   "CH-ENV-CH-ACT" : Bool AT %I76.0, 1 s
   "CH-ENV-CH-TEMP" : Bool AT %I76.1, 1 s
   "CH-ENV-CH-TERM" : Bool AT %I76.2, 1 s
   "CH-ENV-CH-RUN" : Bool AT %I76.3, 1 s
   "BombaTorreON2" : Bool AT %M69.3, 1 s
   "HabV001(1)" : Bool AT %DB90.DBX7.6, 1 s
   "HabV002(1)" : Bool AT %DB90.DBX7.7, 1 s
   "HabV003(1)" : Bool AT %DB90.DBX8.0, 1 s
   "HabV4" : Bool AT %DB90.DBX8.1, 1 s
   "MarchaV001(1)" : Bool AT %DB90.DBX11.0, 1 s
   "MarchaV002(1)" : Bool AT %DB90.DBX11.1, 1 s
   "MarchaV003(1)" : Bool AT %DB90.DBX11.2, 1 s
   "ParadaV001(1)" : Bool AT %DB90.DBX12.5, 1 s
   "ParadaV002(1)" : Bool AT %DB90.DBX12.6, 1 s
   "ParadaV003(1)" : Bool AT %DB90.DBX12.7, 1 s
   "AnimaMenuV001" : Int AT %DB46.DBW24, 1 s
   "AnimaMenuV002" : Int AT %DB46.DBW26, 1 s
   "AnimaMenuV003" : Int AT %DB46.DBW28, 1 s
   "DeshV001" : Bool AT %DB90.DBX9.3, 1 s
   "DeshV002" : Bool AT %DB90.DBX9.4, 1 s
   "DeshV003" : Bool AT %DB90.DBX9.5, 1 s

HMI tags "CompBajaMTA"
   "HabilitaciónMC060" : Bool AT %DB74.DBX3.0, 1 s
   "HabilitaciónMC061" : Bool AT %DB74.DBX3.1, 1 s
   "HabilitaciónMC062" : Bool AT %DB74.DBX3.2, 1 s
   "HabilitaciónMC063" : Bool AT %DB74.DBX3.3, 1 s
   "HabilitaciónMC064" : Bool AT %DB74.DBX3.4, 1 s
   "HabilitaciónMC065" : Bool AT %DB74.DBX3.5, 1 s
   "DeshabilitaciónMC060" : Bool AT %DB74.DBX3.6, 1 s
   "DeshabilitaciónMC061" : Bool AT %DB74.DBX3.7, 1 s
   "DeshabilitaciónMC062" : Bool AT %DB74.DBX4.0, 1 s
   "DeshabilitaciónMC063" : Bool AT %DB74.DBX4.1, 1 s
   "DeshabilitaciónMC064" : Bool AT %DB74.DBX4.2, 1 s
   "DeshabilitaciónMC065" : Bool AT %DB74.DBX4.3, 1 s
   "MarchaMC060" : Bool AT %DB74.DBX4.4, 1 s
   "MarchaMC061" : Bool AT %DB74.DBX4.5, 1 s
   "MarchaMC062" : Bool AT %DB74.DBX4.6, 1 s
   "MarchaMC063" : Bool AT %DB74.DBX4.7, 1 s
   "MarchaMC064" : Bool AT %DB74.DBX5.0, 1 s
   "MarchaMC065" : Bool AT %DB74.DBX5.1, 1 s
   "ParadaMC060" : Bool AT %DB74.DBX5.2, 1 s
   "ParadaMC061" : Bool AT %DB74.DBX5.3, 1 s
   "ParadaMC062" : Bool AT %DB74.DBX5.4, 1 s
   "ParadaMC063" : Bool AT %DB74.DBX5.5, 1 s
   "ParadaMC064" : Bool AT %DB74.DBX5.6, 1 s
   "ParadaMC065" : Bool AT %DB74.DBX5.7, 1 s
   "AnimaMC060" : Byte AT %DB74.DBB9, 1 s
   "AnimaMC061" : Byte AT %DB74.DBB10, 1 s
   "AnimaMC062" : Byte AT %DB74.DBB11, 1 s
   "AnimaMC063" : Byte AT %DB74.DBB12, 1 s
   "AnimaMC064" : Byte AT %DB74.DBB13, 1 s
   "AnimaMC065" : Byte AT %DB74.DBB14, 1 s
   "VerMC060" : Bool, internal
   "VerMC061" : Bool, internal
   "VerMC062" : Bool, internal
   "VerMC063" : Bool, internal
   "VerMC064" : Bool, internal
   "MantM060" : Bool AT %DB74.DBX16.4, 1 s
   "MantM061" : Bool AT %DB74.DBX16.5, 1 s
   "MantM062" : Bool AT %DB74.DBX16.6, 1 s
   "MantM063" : Bool AT %DB74.DBX16.7, 1 s
   "MantM064" : Bool AT %DB74.DBX17.0, 1 s
   "AutoMC060" : Bool AT %DB93.DBX0.0, 1 s
   "AutoMC061" : Bool AT %DB93.DBX0.1, 1 s
   "AutoMC062" : Bool AT %DB93.DBX0.2, 1 s
   "AutoMC063" : Bool AT %DB93.DBX0.3, 1 s
   "AutoMC064" : Bool AT %DB93.DBX0.4, 1 s
   "SponMC060" : Real AT %DB93.DBD2, 1 s
   "SponMC061" : Real AT %DB93.DBD6, 1 s
   "SponMC062" : Real AT %DB93.DBD10, 1 s
   "SponMC063" : Real AT %DB93.DBD14, 1 s
   "SponMC064" : Real AT %DB93.DBD18, 1 s
   "SpoffMC060" : Real AT %DB93.DBD22, 1 s
   "SpoffMC061" : Real AT %DB93.DBD26, 1 s
   "SpoffMC062" : Real AT %DB93.DBD30, 1 s
   "SpoffMC063" : Real AT %DB93.DBD34, 1 s
   "SpoffMC064" : Real AT %DB93.DBD38, 1 s
   "AnimMenuMC060" : Int AT %DB93.DBW44, 1 s
   "AnimMenuMC061" : Int AT %DB93.DBW46, 1 s
   "AnimMenuMC062" : Int AT %DB93.DBW48, 1 s
   "AnimMenuMC063" : Int AT %DB93.DBW50, 1 s
   "AnimMenuMC064" : Int AT %DB93.DBW52, 1 s
   "HabilitarMC060" : Bool AT %M900.0, 1 s
   "AnularSirenaCav" : Bool AT %M600.0, 1 s
   "VerMC65" : Bool, internal

HMI tags "CompresoresAltaMTA"
   "Sop1" : Bool AT %DB124.DBX0.0, 1 s
   "Sop2" : Bool AT %DB124.DBX0.1, 1 s
   "Sop3" : Bool AT %DB124.DBX0.2, 1 s
   "ReqSop1" : Int AT %DB124.DBW8, 1 s
   "ReqSop2" : Int AT %DB124.DBW10, 1 s
   "ReqSop3" : Int AT %DB124.DBW12, 1 s
   "NinSop" : Bool AT %DB124.DBX6.0, 1 s
   "VCMP1" : Int AT %DB125.DBW2, 1 s
   "VCMP2" : Int AT %DB125.DBW4, 1 s
   "VCMP3" : Int AT %DB125.DBW6, 1 s
   "VCMP4" : Int AT %DB125.DBW8, 1 s
   "VCMP5" : Int AT %DB125.DBW10, 1 s
   "IncP1" : Bool AT %DB125.DBX15.4, 100 ms
   "IncP2" : Bool AT %DB125.DBX15.5, 100 ms
   "IncP3" : Bool AT %DB125.DBX15.6, 100 ms
   "IncP4" : Bool AT %DB125.DBX15.7, 100 ms
   "IncP5" : Bool AT %DB125.DBX16.0, 100 ms
   "DecP1" : Bool AT %DB125.DBX16.2, 1 s
   "DecP2" : Bool AT %DB125.DBX16.3, 1 s
   "DecP3" : Bool AT %DB125.DBX16.4, 1 s
   "DecP4" : Bool AT %DB125.DBX16.5, 1 s
   "DecP5" : Bool AT %DB125.DBX16.6, 1 s
   "PriRealCMP1" : Int AT %DB121.DBW16, 1 s
   "PriRealCMP2" : Int AT %DB121.DBW20, 1 s
   "PriRealCMP3" : Int AT %DB121.DBW24, 1 s
   "PriRealCMP4" : Int AT %DB121.DBW28, 1 s
   "PriRealCMP5" : Int AT %DB121.DBW32, 1 s
   "Auto1" : Bool AT %DB88.DBX10.0, 1 s
   "Auto2" : Bool AT %DB88.DBX10.1, 1 s
   "Auto3" : Bool AT %DB88.DBX10.2, 1 s
   "Auto4" : Bool AT %DB88.DBX10.3, 1 s
   "Auto5" : Bool AT %DB88.DBX10.4, 1 s
   "IndV1" : Bool AT %DB121.DBX1.5, 100 ms
   "IndV2" : Bool AT %DB121.DBX1.6, 100 ms
   "IndV3" : Bool AT %DB121.DBX1.7, 100 ms
   "IndV4" : Bool AT %DB121.DBX2.0, 100 ms
   "IndV5" : Bool AT %DB121.DBX2.1, 100 ms
   "IndR1" : Bool AT %DB121.DBX2.3, 100 ms
   "IndR2" : Bool AT %DB121.DBX2.4, 100 ms
   "IndR3" : Bool AT %DB121.DBX2.5, 100 ms
   "IndR4" : Bool AT %DB121.DBX2.6, 100 ms
   "IndR5" : Bool AT %DB121.DBX2.7, 100 ms
   "Est1" : Word AT %DB120.DBW0, 1 s
   "Est2" : Word AT %DB120.DBW2, 1 s
   "Est3" : Word AT %DB120.DBW4, 1 s
   "Est4" : Word AT %DB120.DBW6, 1 s
   "Est5" : Word AT %DB120.DBW8, 1 s
   "LimSUP1" : Real AT %DB122.DBD0, 1 s
   "LimSUP2" : Real AT %DB122.DBD4, 1 s
   "LimSUP3" : Real AT %DB122.DBD8, 1 s
   "LimSUP4" : Real AT %DB122.DBD12, 1 s
   "LimSUP5" : Real AT %DB122.DBD16, 1 s
   "LimINF1" : Real AT %DB122.DBD24, 1 s
   "LimINF2" : Real AT %DB122.DBD28, 1 s
   "LimINF3" : Real AT %DB122.DBD32, 1 s
   "LimINF4" : Real AT %DB122.DBD36, 1 s
   "LimINF5" : Real AT %DB122.DBD40, 1 s
   "PresMaX" : Real AT %DB122.DBD56, 1 s
   "Delta" : Real AT %DB122.DBD48, 1 s
   "Hist" : Real AT %DB122.DBD52, 1 s
   "CompReq" : Int AT %DB121.DBW4, 1 s
   "CompReqINI" : Int AT %DB124.DBW14, 1 s
   "AnimMenuMC001" : Int AT %DB135.DBW0, 1 s
   "AnimMenuMC002" : Int AT %DB135.DBW2, 1 s
   "AnimMenuMC003" : Int AT %DB135.DBW4, 1 s
   "AnimMenuMC004" : Int AT %DB135.DBW6, 1 s
   "AnimMenuMC005" : Int AT %DB135.DBW8, 1 s
   "SPON1" : Real AT %DB135.DBD12, 1 s
   "SPON2" : Real AT %DB135.DBD16, 1 s
   "SPON3" : Real AT %DB135.DBD20, 1 s
   "SPON4" : Real AT %DB135.DBD24, 1 s
   "SPON5" : Real AT %DB135.DBD28, 1 s
   "SPOFF1" : Real AT %DB135.DBD36, 1 s
   "SPOFF2" : Real AT %DB135.DBD40, 1 s
   "SPOFF3" : Real AT %DB135.DBD44, 1 s
   "SPOFF4" : Real AT %DB135.DBD48, 1 s
   "SPOFF5" : Real AT %DB135.DBD52, 1 s
   "MantMC001" : Bool AT %DB135.DBX60.0, 1 s
   "MantMC002" : Bool AT %DB135.DBX60.1, 1 s
   "MantMC003" : Bool AT %DB135.DBX60.2, 1 s
   "MantMC004" : Bool AT %DB135.DBX60.3, 1 s
   "MantMC005" : Bool AT %DB135.DBX60.4, 1 s
   "IndVparp1" : Bool AT %DB121.DBX70.0, 1 s
   "IndVparp2" : Bool AT %DB121.DBX70.1, 1 s
   "IndVparp3" : Bool AT %DB121.DBX70.2, 1 s
   "IndVparp4" : Bool AT %DB121.DBX70.3, 1 s
   "IndVparp5" : Bool AT %DB121.DBX70.4, 1 s
   "TiempoenVacío" : Int AT %DB123.DBW4, 1 s
   "TiemposinReq" : Int AT %DB123.DBW10, 1 s
   "TiempoSop" : Int AT %DB124.DBW4, 1 s
   "HistCRT" : Real AT %DB122.DBD60, 1 s
   "LimINFCRT" : Real AT %DB122.DBD68, 1 s
   "LimSUPCRT" : Real AT %DB122.DBD64, 1 s
   "PanMCH1" : Bool AT %DB88.DBX6.0, 1 s
   "PanMCH2" : Bool AT %DB88.DBX6.1, 1 s
   "PanMCH3" : Bool AT %DB88.DBX6.2, 1 s
   "PanMCH4" : Bool AT %DB88.DBX6.3, 1 s
   "PanMCH5" : Bool AT %DB88.DBX6.4, 1 s
   "MarchaMC001" : Bool AT %DB135.DBX61.4, 1 s
   "MarchaMC002" : Bool AT %DB135.DBX61.5, 1 s
   "MarchaMC003" : Bool AT %DB135.DBX61.6, 1 s
   "MarchaMC004" : Bool AT %DB135.DBX61.7, 1 s
   "MarchaMC005" : Bool AT %DB135.DBX62.0, 1 s
   "ParadaMC001" : Bool AT %DB135.DBX62.2, 1 s
   "ParadaMC002" : Bool AT %DB135.DBX62.3, 1 s
   "ParadaMC003" : Bool AT %DB135.DBX62.4, 1 s
   "ParadaMC004" : Bool AT %DB135.DBX62.5, 1 s
   "ParadaMC005" : Bool AT %DB135.DBX62.6, 1 s
   "AnimMotorMC001" : Byte AT %DB46.DBB40, 1 s
   "AnimMotorMC002" : Byte AT %DB46.DBB41, 1 s
   "AnimMotorMC003" : Byte AT %DB46.DBB42, 1 s
   "AnimMotorMC004" : Byte AT %DB46.DBB43, 1 s
   "AnimMotorMC005" : Byte AT %DB46.DBB44, 1 s
   "EV1" : Bool AT %Q2.0, 1 s
   "EV2" : Bool AT %Q2.1, 1 s
   "EV3" : Bool AT %Q2.2, 1 s
   "EV4" : Bool AT %Q2.3, 1 s
   "EV5" : Bool AT %Q2.4, 1 s
   "HORAS1" : DInt AT %DB73.DBD0, 1 s
   "HORAS2" : DInt AT %DB73.DBD4, 1 s
   "HORAS3" : DInt AT %DB73.DBD8, 1 s
   "HORAS4" : DInt AT %DB73.DBD12, 1 s
   "HORAS5" : DInt AT %DB73.DBD16, 1 s
   "MIN1" : Int AT %DB73.DBW24, 1 s
   "MIN2" : Int AT %DB73.DBW26, 1 s
   "MIN3" : Int AT %DB73.DBW28, 1 s
   "MIN4" : Int AT %DB73.DBW30, 1 s
   "MIN5" : Int AT %DB73.DBW32, 1 s
   "MarchaOK1" : Bool AT %DB135.DBX60.6, 1 s
   "MarchaOK2" : Bool AT %DB135.DBX60.7, 1 s
   "MarchaOK3" : Bool AT %DB135.DBX61.0, 1 s
   "MarchaOK4" : Bool AT %DB135.DBX61.1, 1 s
   "MarchaOK5" : Bool AT %DB135.DBX61.2, 1 s
   "ForzarMarcha1" : Bool AT %DB136.DBX0.0, 1 s
   "ForzarMarcha2" : Bool AT %DB136.DBX0.1, 1 s
   "ForzarMarcha3" : Bool AT %DB136.DBX0.2, 1 s
   "ForzarMarcha4" : Bool AT %DB136.DBX0.3, 1 s
   "ForzarMarcha5" : Bool AT %DB136.DBX0.4, 1 s
   "ForzarParada1" : Bool AT %DB136.DBX0.6, 1 s
   "ForzarParada2" : Bool AT %DB136.DBX0.7, 1 s
   "ForzarParada3" : Bool AT %DB136.DBX1.0, 1 s
   "ForzarParada4" : Bool AT %DB136.DBX1.1, 1 s
   "ForzarParada5" : Bool AT %DB136.DBX1.2, 1 s
   "SPONF1" : Real AT %DB136.DBD4, 1 s
   "SPONF2" : Real AT %DB136.DBD8, 1 s
   "SPONF3" : Real AT %DB136.DBD12, 1 s
   "SPONF4" : Real AT %DB136.DBD16, 1 s
   "SPONF5" : Real AT %DB136.DBD20, 1 s
   "SPOFFF1" : Real AT %DB136.DBD28, 1 s
   "SPOFFF2" : Real AT %DB136.DBD32, 1 s
   "SPOFFF3" : Real AT %DB136.DBD36, 1 s
   "SPOFFF4" : Real AT %DB136.DBD40, 1 s
   "SPOFFF5" : Real AT %DB136.DBD44, 1 s
   "ForzandoMarcha1" : Bool AT %DB136.DBX1.4, 1 s
   "ForzandoMarcha2" : Bool AT %DB136.DBX1.5, 1 s
   "ForzandoMarcha3" : Bool AT %DB136.DBX1.6, 1 s
   "ForzandoMarcha4" : Bool AT %DB136.DBX1.7, 1 s
   "ForzandoMarcha5" : Bool AT %DB136.DBX2.0, 1 s
   "MediaCargaBellis" : Bool AT %DB135.DBX63.0, 1 s
   "SPONF3b" : Real AT %DB136.DBD52, 1 s
   "SPOFFF3b" : Real AT %DB136.DBD56, 1 s
   "EV3b" : Bool AT %Q3.2, 1 s
   "TiempoMaxBellismedia" : Int AT %DB63.DBW4, 1 s
   "Est6" : Int AT %DB120.DBW10, 1 s
   "PriRealCMP6" : Int AT %DB121.DBW36, 1 s
   "IndV6" : Bool AT %DB121.DBX2.2, 1 s

HMI tags "IluminaciónMTA"
   "TiempoIluminación" : Word AT %DB87.DBW0, 1 s
   "EncendidoPanel" : Bool AT %DB87.DBX2.0, 1 s
   "ApagadoPanel" : Bool AT %DB87.DBX2.1, 1 s
   "ON" : Bool AT %DB87.DBX2.2, 1 s
   "MantenerON" : Bool AT %DB87.DBX2.3, 1 s
   "AlarmaBoosters" : Bool AT %M330.4, 1 s

HMI tags "SecadoresAltaMTA"
   "AnimaMS050" : Byte AT %DB81.DBB6, 1 s
   "AnimaMS051" : Byte AT %DB81.DBB7, 1 s
   "AnimaMS052" : Byte AT %DB81.DBB8, 1 s
   "AnimaMS053" : Byte AT %DB81.DBB9, 1 s
   "DeshabilitaciónMS050" : Bool AT %DB81.DBX2.4, 1 s
   "DeshabilitaciónMS051" : Bool AT %DB81.DBX2.5, 1 s
   "DeshabilitaciónMS052" : Bool AT %DB81.DBX2.6, 1 s
   "DeshabilitaciónMS053" : Bool AT %DB81.DBX2.7, 1 s
   "HabilitaciónMS050" : Bool AT %DB81.DBX2.0, 1 s
   "HabilitaciónMS051" : Bool AT %DB81.DBX2.1, 1 s
   "HabilitaciónMS052" : Bool AT %DB81.DBX2.2, 1 s
   "HabilitaciónMS053" : Bool AT %DB81.DBX2.3, 1 s
   "MantMS050" : Bool AT %DB81.DBX11.0, 1 s
   "MantMS051" : Bool AT %DB81.DBX11.1, 1 s
   "MantMS052" : Bool AT %DB81.DBX11.2, 1 s
   "MantMS053" : Bool AT %DB81.DBX11.3, 1 s
   "MarchaMS050" : Bool AT %DB81.DBX3.0, 1 s
   "MarchaMS051" : Bool AT %DB81.DBX3.1, 1 s
   "MarchaMS052" : Bool AT %DB81.DBX3.2, 1 s
   "MarchaMS053" : Bool AT %DB81.DBX3.3, 1 s
   "ParadaMS050" : Bool AT %DB81.DBX3.4, 1 s
   "ParadaMS051" : Bool AT %DB81.DBX3.5, 1 s
   "ParadaMS052" : Bool AT %DB81.DBX3.6, 1 s
   "ParadaMS053" : Bool AT %DB81.DBX3.7, 1 s
   "AnimaMenuMS050" : Int AT %DB46.DBW14, 1 s
   "AnimaMenuMS051" : Int AT %DB46.DBW16, 1 s
   "AnimaMenuMS052" : Int AT %DB46.DBW18, 1 s
   "AnimaMenuMS053" : Int AT %DB46.DBW20, 1 s
   "Enc1MS050" : Int AT %DB81.DBW12, 1 s
   "Enc2MS050" : Int AT %DB81.DBW14, 1 s
   "Enc1MS051" : Int AT %DB81.DBW16, 1 s
   "Enc2MS051" : Int AT %DB81.DBW18, 1 s
   "Enc1MS052" : Int AT %DB81.DBW20, 1 s
   "Enc2MS052" : Int AT %DB81.DBW22, 1 s
   "Enc1MS053" : Int AT %DB81.DBW24, 1 s
   "Enc2MS053" : Int AT %DB81.DBW26, 1 s
   "AutoMS050" : Bool AT %DB81.DBX28.0, 1 s
   "AutoMS051" : Bool AT %DB81.DBX28.1, 1 s
   "AutoMS052" : Bool AT %DB81.DBX28.2, 1 s
   "AutoMS053" : Bool AT %DB81.DBX28.3, 1 s

HMI tags "SecadoresBaja"
   "AnimaMS054" : Byte AT %DB46.DBB30, 1 s
   "AnimaMS055" : Byte AT %DB46.DBB31, 1 s
   "DeshabilitaciónMS054" : Bool AT %DB49.DBX1.2, 1 s
   "DeshabilitaciónMS055" : Bool AT %DB49.DBX1.3, 1 s
   "HabilitaciónMS054" : Bool AT %DB49.DBX1.0, 1 s
   "HabilitaciónMS055" : Bool AT %DB49.DBX1.1, 1 s
   "MarchaMS054" : Bool AT %DB49.DBX1.4, 1 s
   "MarchaMS055" : Bool AT %DB49.DBX1.5, 1 s
   "ParadaMS054" : Bool AT %DB49.DBX1.6, 1 s
   "ParadaMS055" : Bool AT %DB49.DBX1.7, 1 s
   "MantMS054" : Bool AT %DB49.DBX5.4, 1 s
   "MantMS055" : Bool AT %DB49.DBX5.5, 1 s

HMI tags "SENTRON PAC 3200"
   "Tension Fase R" : Float AT %MW1, 1 s
   "Tension fase S" : Float AT %MW3, 1 s
   "Tension Fase T" : Float AT %MW5, 1 s
   "Tension Linea RS" : Float AT %MW7, 1 s
   "Tension Linea ST" : Float AT %MW9, 1 s
   "Tension Linea TR" : Float AT %MW11, 1 s
   "Corriente fase R" : Float AT %MW13, 1 s
   "Corriente Fase S" : Float AT %MW15, 1 s
   "Corriente Fase T" : Float AT %MW17, 1 s
   "Pot.Apa R" : Float AT %MW19, 1 s
   "Pot.Apa S" : Float AT %MW21, 1 s
   "Pot.Apa T" : Float AT %MW23, 1 s
   "Pot.Act R" : Float AT %MW25, 1 s
   "Pot.Act S" : Float AT %MW27, 1 s
   "Pot.Act T" : Float AT %MW29, 1 s
   "Pot.ReAct R" : Float AT %MW31, 1 s
   "Pot.ReAct S" : Float AT %MW33, 1 s
   "Pot.ReAct T" : Float AT %MW35, 1 s
   "Coseno R" : Float AT %MW37, 1 s
   "Coseno S" : Float AT %MW39, 1 s
   "Coseno T" : Float AT %MW41, 1 s
   "THD-R TensionFase R" : Float AT %MW43, 1 s
   "THD-R Tension Fase S" : Float AT %MW45, 1 s
   "THD-R Tension Fase T" : Float AT %MW47, 1 s
   "THD-R Corriente Fase R" : Float AT %MW49, 1 s
   "THD-R Corriente Fase S" : Float AT %MW51, 1 s
   "THD-R Corriente Fase T" : Float AT %MW53, 1 s
   "Frecuencia" : Float AT %MW55, 1 s
   "Tension Media Fase" : Float AT %MW57, 1 s
   "Tension Media de Linea" : Float AT %MW59, 1 s
   "Corriente Media" : Float AT %MW61, 1 s
   "Pot Apa Total" : Float AT %MW63, 1 s
   "Pot Act Total" : Float AT %MW65, 1 s
   "Pot ReAct Total" : Float AT %MW67, 1 s
   "coseno Total" : Float AT %MW69, 1 s
   "desbalance de tension" : Float AT %MW71, 1 s
   "desbalance de corriente" : Float AT %MW73, 1 s
   "Tension Maxima R" : Float AT %MW75, 1 s
   "Tension Maxima S" : Float AT %MW77, 1 s
   "Tension Maxima T" : Float AT %MW79, 1 s
   "Tension Maxima RS" : Float AT %MW81, 1 s
   "Tension Maxima ST" : Float AT %MW83, 1 s
   "Tension Maxima TR" : Float AT %MW85, 1 s
   "Corriente Maxima R" : Float AT %MW87, 1 s
   "Corriente Maxima S" : Float AT %MW89, 1 s
   "Corriente Maxima T" : Float AT %MW91, 1 s

HMI tags "TorresCav-MTA"
   "AnimaMV030" : Byte AT %DB46.DBB36, 1 s
   "AnimaMV031" : Byte AT %DB46.DBB37, 1 s
   "AnimaMP014" : Byte AT %DB46.DBB38, 1 s
   "AnimaMP015" : Byte AT %DB46.DBB39, 1 s
   "DeshabilitaciónMV030" : Bool AT %DB21.DBX2.4, 1 s
   "DeshabilitaciónMV031" : Bool AT %DB21.DBX2.5, 1 s
   "DeshabilitaciónMP014" : Bool AT %DB21.DBX2.6, 1 s
   "DeshabilitaciónMP015" : Bool AT %DB21.DBX2.7, 1 s
   "HabilitaciónMV030" : Bool AT %DB21.DBX2.0, 1 s
   "HabilitaciónMV031" : Bool AT %DB21.DBX2.1, 1 s
   "HabilitaciónMP014" : Bool AT %DB21.DBX2.2, 1 s
   "HabilitaciónMP015" : Bool AT %DB21.DBX2.3, 1 s
   "MantMV030" : Bool AT %DB21.DBX10.0, 1 s
   "MantMV031" : Bool AT %DB21.DBX10.1, 1 s
   "MantMP014" : Bool AT %DB21.DBX10.2, 1 s
   "MantMP015" : Bool AT %DB21.DBX10.3, 1 s
   "MarchaMV030" : Bool AT %DB21.DBX3.0, 1 s
   "MarchaMV031" : Bool AT %DB21.DBX3.1, 1 s
   "MarchaMP014" : Bool AT %DB21.DBX3.2, 1 s
   "MarchaMP015" : Bool AT %DB21.DBX3.3, 1 s
   "ParadaMV030" : Bool AT %DB21.DBX3.4, 1 s
   "ParadaMV031" : Bool AT %DB21.DBX3.5, 1 s
   "ParadaMP014" : Bool AT %DB21.DBX3.6, 1 s
   "ParadaMP015" : Bool AT %DB21.DBX3.7, 1 s
   "MenuV030" : Int AT %DB46.DBW32, 1 s
   "MenuV031" : Int AT %DB46.DBW34, 1 s

discrete alarms
   1: 'Falla Conexión con sensor de Temperatura torres de Cavaleto', class MTA, trigger "Rec13" bit 9
   2: 'Falla Conexión con sensor de Temperatura torres de Chillers', class MTA, trigger "Rec13" bit 10
   3: 'Falla Conexión con sensor de Presión de ALTA', class MTA, trigger "Rec13" bit 11
   4: 'Falla Conexión con sensor de Presión de ALTA redundante', class MTA, trigger "Rec13" bit 12
   5: 'Falla Conexión con sensor de Presión de Baja', class MTA, trigger "Rec13" bit 13
   6: 'Falla Presión de Alta en Límite Mínimo', class MTA, trigger "Rec13" bit 14
   7: 'Falla Presión de Alta en demasiado Baja', class MTA, trigger "Rec13" bit 15
   8: 'Falla Presión de Alta en demasiado Alta', class MTA, trigger "Rec14" bit 8
   9: 'Falla Presión de Alta en Límite Máximo', class MTA, trigger "Rec14" bit 9
   10: 'Falla Presión de Baja en Límite Mínimo', class MTA, trigger "Rec14" bit 10
   11: 'Falla Presión de Baja en demasiado Baja', class MTA, trigger "Rec14" bit 11
   12: 'Falla Presión de Baja en demasiado Alta', class MTA, trigger "Rec14" bit 12
   13: 'Falla Contactor - MS050 - Secador de Alta ABC1', class MTA, trigger "Rec6" bit 8
   14: 'Falla Guardamotor - MS051 - Secador de Alta ABC3', class MTA, trigger "Rec6" bit 9
   15: 'Falla Presión de Baja en Límite Máximo', class MTA, trigger "Rec14" bit 13
   16: 'Falla en chiller de envasado chico', class MTA, trigger "Rec14" bit 14
   17: 'Falla en chiller de soplado chico', class MTA, trigger "Rec14" bit 15
   18: 'El Compresor ABC2 alcanzó la máxima cantidad de horas sin mantenimiento #1', class MTA, trigger "Rec15" bit 8
   19: 'El Compresor ABC3 alcanzó la máxima cantidad de horas sin mantenimiento #1', class MTA, trigger "Rec15" bit 9
   20: 'El Compresor Bellis alcanzó la máxima cantidad de horas sin mantenimiento #1', class MTA, trigger "Rec15" bit 10
   21: 'El Compresor ABC4 alcanzó la máxima cantidad de horas sin mantenimiento #1', class MTA, trigger "Rec15" bit 11
   22: 'El Compresor ABC5 alcanzó la máxima cantidad de horas sin mantenimiento #1', class MTA, trigger "Rec15" bit 12
   23: 'Falla algún contactor en Booster 1', class MTA, trigger "Rec15" bit 13
   24: 'Falla algún guardamotor en Booster 1', class MTA, trigger "Rec15" bit 14
   25: 'Presión Alta en Booster', class MTA, trigger "Rec15" bit 15
   26: 'Falla algún contactor en Booster 2', class MTA, trigger "Rec16" bit 8
   27: 'Falla algún guardamotor en Booster 2', class MTA, trigger "Rec16" bit 9
   28: 'Error lectura analógica Presión Boosters', class MTA, trigger "Rec16" bit 10
   29: 'Bombas Torres de Agua Cavaleto detenidas por falla en Flujostato', class MTA, trigger "Rec16" bit 11
   30: 'Ventiladores Torres de Agua Cavaleto detenidas por falla en Flujostato', class MTA, trigger "Rec16" bit 12
   31: 'Ninguna Bomba Torres de Agua Cabaleto en Marcha', class MTA, trigger "Rec16" bit 13
   32: 'Compresores Alta Detenidos por Flujostato Torres de Agua Cabaleto', class MTA, trigger "Rec16" bit 14
   33: 'Compresores Alta Detenidos por Ninguna Bomba en Marcha en Torres de Agua Cabaleto', class MTA, trigger "Rec16" bit 15
   50: 'Falla Contactor - MS051 - Secador de Alta ABC3', class MTA, trigger "Rec6" bit 10
   53: 'Falla Guardamotor - MS052 - Secador de Alta ABC2', class MTA, trigger "Rec6" bit 11
   66: 'Falla Guardamotor MS054 - Secador de Baja SULLAIR 1', class MTA, trigger "Rec7" bit 8
   67: 'Falla Contactor MS054 - Secador de Baja SULLAIR 1', class MTA, trigger "Rec7" bit 9
   68: 'Falla Guardamotor MS055 - Secador de Baja SULLAIR 2', class MTA, trigger "Rec7" bit 10
   69: 'Falla Contactor MS055 - Secador de Baja SULLAIR 2', class MTA, trigger "Rec7" bit 11
   70: 'Falla Guardamotor - MV030 - Ventilador 2 Torres de enfriamiento Cavaleto', class MTA, trigger "Rec7" bit 12
   71: 'Falla Contactor - MV030 - Ventilador 2 Torres de enfriamiento Cavaleto', class MTA, trigger "Rec7" bit 13
   72: 'Falla Guardamotor - MV031 - Ventilador 1 Torres de enfriamiento Cavaleto', class MTA, trigger "Rec7" bit 14
   73: 'Falla Contactor - MV031 - Ventilador 1 Torres de enfriamiento Cavaleto', class MTA, trigger "Rec7" bit 15
   74: 'Falla Guardamotor - MP014 - Bomba 1 Torres de enfriamiento Cavaleto', class MTA, trigger "Rec8" bit 8
   75: 'Falla Contactor - MP014 - Bomba 1 Torres de enfriamiento Cavaleto', class MTA, trigger "Rec8" bit 9
   76: 'Falla Guardamotor - MP015 - Bomba 2 Torres de enfriamiento Cavaleto', class MTA, trigger "Rec8" bit 10
   77: 'Falla Contactor - MP015 - Bomba 2 Torres de enfriamiento Cavaleto', class MTA, trigger "Rec8" bit 11
   78: 'Falla Guardamotor - MC001 - Compresor de Alta ABC2', class MTA, trigger "Rec8" bit 12
   79: 'Falla Contactor - MC001 - Compresor de Alta ABC2', class MTA, trigger "Rec8" bit 13
   80: 'Falla Guardamotor - MC002 - Compresor de Alta ABC3', class MTA, trigger "Rec8" bit 14
   81: 'Falla Contactor - MC002 - Compresor de Alta ABC3', class MTA, trigger "Rec8" bit 15
   82: 'Falla Guardamotor - MC003 - Compresor de Alta BELLIS', class MTA, trigger "Rec9" bit 8
   83: 'Falla Contactor - MC003 - Compresor de Alta BELLIS', class MTA, trigger "Rec9" bit 9
   87: 'Falla Contactor - MS052 - Secador de Alta ABC2', class MTA, trigger "Rec6" bit 12
   88: 'Falla Guardamotor - MS053 - Secador de Alta FARGON', class MTA, trigger "Rec6" bit 13
   89: 'Falla Contactor - MS053 - Secador de Alta FARGON', class MTA, trigger "Rec6" bit 14
   90: 'Falla Presostato Chillers', class MTA, trigger "Rec6" bit 15
   91: 'Falla Guardamotor - MC004 - Compresor de Alta ABC4', class MTA, trigger "Rec9" bit 10
   92: 'Falla Contactor - MC004 - Compresor de Alta ABC4', class MTA, trigger "Rec9" bit 11
   93: 'Falla Guardamotor - MC005 - Compresor de Alta ABC5', class MTA, trigger "Rec9" bit 12
   94: 'Falla Contactor - MC005 - Compresor de Alta ABC5', class MTA, trigger "Rec9" bit 13
   95: 'Falla Flujostato Torres Caveleto', class MTA, trigger "Rec9" bit 14
   96: 'Falla Compresor ABC2 Baja Presion de Aceite', class MTA, trigger "Rec9" bit 15
   97: 'Falla Compresor ABC2 Baja Presion de Agua', class MTA, trigger "Rec10" bit 8
   98: 'Falla Compresor ABC2 Alta Temperatura de Aire', class MTA, trigger "Rec10" bit 9
   99: 'Falla Compresor ABC2 Alta Temperatura de agua', class MTA, trigger "Rec10" bit 10
   100: 'Falla Compresor ABC3 Baja Presion de Aceite', class MTA, trigger "Rec10" bit 11
   101: 'Falla Compresor ABC3 Baja Presion de Agua', class MTA, trigger "Rec10" bit 12
   102: 'Falla Compresor ABC3 Alta Temperatura de Aire', class MTA, trigger "Rec10" bit 13
   103: 'Falla Compresor ABC3 Alta Temperatura de agua', class MTA, trigger "Rec10" bit 14
   104: 'Falla Compresor ABC4 Baja Presion de Aceite', class MTA, trigger "Rec10" bit 15
   105: 'Falla Compresor ABC4 Alta Temperatura de Aire', class MTA, trigger "Rec11" bit 8
   106: 'Falla Compresor ABC4 Alta Temperatura de Aire', class MTA, trigger "Rec11" bit 9
   107: 'Falla Compresor ABC4 Alta Temperatura de agua', class MTA, trigger "Rec11" bit 10
   108: 'Falla Compresor ABC5 Baja Presion de Aceite', class MTA, trigger "Rec11" bit 11
   109: 'Falla Compresor ABC5 Alta Temperatura de Aire', class MTA, trigger "Rec11" bit 12
   110: 'Falla Compresor ABC5 Alta Temperatura de Aire', class MTA, trigger "Rec11" bit 13
   111: 'Falla Compresor ABC5 Alta Temperatura de agua', class MTA, trigger "Rec11" bit 14
   112: 'Falla Compresor Bellis & MHW28 Baja Presion Aceite', class MTA, trigger "Rec11" bit 15
   113: 'Falla Compresor Bellis & MHW28 Baja Presion de Agua', class MTA, trigger "Rec12" bit 8
   114: 'Falla Compresor Bellis & MHW28 Alta temperatura de Aire', class MTA, trigger "Rec12" bit 9
   115: 'Falla Compresor Bellis & MHW28 Alta temperatura de Agua', class MTA, trigger "Rec12" bit 10
   116: 'Falla Compresor Bellis & MHW28 Falla de Flujostato', class MTA, trigger "Rec12" bit 11
   117: 'Compresor ABC2 Requiere Marcha', class MTA, trigger "Rec12" bit 12
   118: 'Compresor ABC3 Requiere Marcha', class MTA, trigger "Rec12" bit 13
   119: 'Compresor Bellis Requiere Marcha', class MTA, trigger "Rec12" bit 14
   120: 'Compresor ABC4 Requiere Marcha', class MTA, trigger "Rec12" bit 15
   121: 'Compresor ABC5 Requiere Marcha', class MTA, trigger "Rec13" bit 8
   125: 'Falla Contactor - V001 - Ventilador 1 Torres de enfriamiento Chillers', class MTA, trigger "Rec4" bit 8
   126: 'Falla Guardamotor - V001 - Ventilador 1 Torres de enfriamiento Chillers', class MTA, trigger "Rec3" bit 15
   127: 'Falla Guardamotor - V003 - Ventilador 3 Torres de enfriamiento Chillers', class MTA, trigger "Rec4" bit 11
   128: 'Falla Contactor - V002 - Ventilador 2 Torres de enfriamiento Chillers', class MTA, trigger "Rec4" bit 10
   129: 'Falla Guardamotor - V002 - Ventilador 2 Torres de enfriamiento Chillers', class MTA, trigger "Rec4" bit 9
   130: 'Falla Guardamotor - MP018 - Bomba 1 Torres de enfriamiento Chillers', class MTA, trigger "Rec3" bit 11
   131: 'Falla Contactor - MP013 - Bomba Backup Ch. Envasado', class MTA, trigger "Rec3" bit 10
   132: 'Falla Guardamotor - MP013 - Bomba Backup Ch. Envasado', class MTA, trigger "Rec3" bit 9
   133: 'Falla Contactor - MP019 - Bomba 2 Torres de enfriamiento Chillers', class MTA, trigger "Rec3" bit 14
   134: 'Falla Guardamotor - MP019 - Bomba 2 Torres de enfriamiento Chillers', class MTA, trigger "Rec3" bit 13
   135: 'Falla Contactor - MP018 - Bomba 1 Torres de enfriamiento Chillers', class MTA, trigger "Rec3" bit 12
   136: 'Falla Contactor - V003 - Ventilador 3 Torres de enfriamiento Chillers', class MTA, trigger "Rec4" bit 12
   137: 'Falla Guardamotor - MC061 - Compresor de Baja SULLAIR 1', class MTA, trigger "Rec4" bit 15
   138: 'Falla Contactor - MC060 - Compresor de Baja SULLAIR 2', class MTA, trigger "Rec4" bit 14
   139: 'Falla Guardamotor - MC060 - Compresor de Baja SULLAIR 2', class MTA, trigger "Rec4" bit 13
   140: 'Falla Contactor - MP012 - Bomba Principal Ch. Envasado', class MTA, trigger "Rec3" bit 8
   141: 'Alarma Presente en Chiller de envasado Grande', class MTA, trigger "Rec1" bit 8
   142: 'Alarma Presente en Chiller de soplado Grande', class MTA, trigger "Rec0" bit 15
   143: 'Ningún chiller de envasado habilitado', class MTA, trigger "Rec0" bit 14
   144: 'Falla Guardamotor - MT007 -Sopladora Línea 1', class MTA, trigger "Rec1" bit 11
   145: 'Chiller de envasado Grande en su máxima capacidad', class MTA, trigger "Rec1" bit 10
   146: 'Chiller de soplado Grande en su máxima capacidad', class MTA, trigger "Rec1" bit 9
   147: 'Ninguna bomba de intercambiador de envasado en marcha', class MTA, trigger "Rec0" bit 10
   148: 'Ninguna bomba de chillers de soplado en marcha', class MTA, trigger "Rec0" bit 9
   149: 'Ninguna bomba de intercambiador de soplado en marcha', class MTA, trigger "Rec0" bit 8
   150: 'Ningún Chiller de soplado habilitado', class MTA, trigger "Rec0" bit 13
   151: 'Ninguna bomba de torre de enfiamiento de chillers en marcha', class MTA, trigger "Rec0" bit 12
   152: 'Ninguna bomba de chillers de envasado en marcha', class MTA, trigger "Rec0" bit 11
   153: 'Falla Contactor - MT007 -Sopladora Línea 1', class MTA, trigger "Rec1" bit 12
   154: 'Falla Contactor - MP010 - Bomba Principal Ch. Soplado', class MTA, trigger "Rec2" bit 12
   155: 'Falla Guardamotor - MP010 - Bomba Principal Ch. Soplado', class MTA, trigger "Rec2" bit 11
   156: 'Falla Contactor - MT010 - Bomba Int L1 y Manomec', class MTA, trigger "Rec2" bit 10
   157: 'Falla Guardamotor - MP012 - Bomba Principal Ch. Envasado', class MTA, trigger "Rec2" bit 15
   158: 'Falla Contactor - MP011 - Bomba Backup Ch. Soplado', class MTA, trigger "Rec2" bit 14
   159: 'Falla Guardamotor - MP011 - Bomba Backup Ch. Soplado', class MTA, trigger "Rec2" bit 13
   160: 'Falla Guardamotor - MT009 - Bomba Int. L3 y L5', class MTA, trigger "Rec1" bit 15
   161: 'Falla Contactor - MT008 - Sopladora Línea 3 y Man.', class MTA, trigger "Rec1" bit 14
   162: 'Falla Guardamotor - MT008 - Sopladora Línea 3 y Man.', class MTA, trigger "Rec1" bit 13
   163: 'Falla Guardamotor - MT010 - Bomba Int L1 y Manomec', class MTA, trigger "Rec2" bit 9
   164: 'Falla Contactor - MT009 - Bomba Int. L3 y L5', class MTA, trigger "Rec2" bit 8
   165: 'Falla Contactor - MC061 - Compresor de Baja SULLAIR 1', class MTA, trigger "Rec5" bit 8
   166: 'Falla Guardamotor - MC062 - Compresor de Baja SULLAIR 0', class MTA, trigger "Rec5" bit 9
   167: 'Falla Contactor - MC062 - Compresor de Baja SULLAIR 0', class MTA, trigger "Rec5" bit 10
   168: 'Falla Guardamotor - MC063 - Compresor de Baja ATLAS 3', class MTA, trigger "Rec5" bit 11
   169: 'Falla Contactor - MC063 - Compresor de Baja ATLAS 3', class MTA, trigger "Rec5" bit 12
   170: 'Falla Guardamotor - MC064 - Compresor de Baja ATLAS 2', class MTA, trigger "Rec5" bit 13
   171: 'Falla Contactor - MC064 - Compresor de Baja ATLAS 2', class MTA, trigger "Rec5" bit 14
   172: 'Falla Guardamotor - MS050 - Secador de Alta ABC1', class MTA, trigger "Rec5" bit 15
   34: 'Falla Compresor ABC1 Baja Presion de Aceite', class MTA, trigger "Rec18" bit 8
   35: 'Falla Compresor ABC1 Baja Presión de agua', class MTA, trigger "Rec18" bit 9
   36: 'Falla Compresor ABC1 Alta Temperatura de Aire', class MTA, trigger "Rec18" bit 10
   37: 'Falla Compresor ABC1 Alta Temperatura de agua', class MTA, trigger "Rec18" bit 11
   38: 'Falla Guardamotor - MC006 - Compresor de Alta ABC1', class MTA, trigger "Rec18" bit 12
   39: 'Falla Contactor - MC006 - Compresor de Alta ABC1', class MTA, trigger "Rec18" bit 13
   40: 'Compresor ABC1 Requiere Marcha', class MTA, trigger "Rec18" bit 14
   41: 'El Compresor ABC1 alcanzó la máxima cantidad de horas sin mantenimiento #1', class MTA, trigger "Rec4" bit 15
   42: 'El Compresor ABC2 alcanzó la máxima cantidad de horas sin mantenimiento #2', class MTA, trigger "Rec19" bit 8
   43: 'El Compresor ABC3 alcanzó la máxima cantidad de horas sin mantenimiento #2', class MTA, trigger "Rec19" bit 9
   44: 'El Compresor Bellis alcanzó la máxima cantidad de horas sin mantenimiento #2', class MTA, trigger "Rec19" bit 10
   45: 'El Compresor ABC4 alcanzó la máxima cantidad de horas sin mantenimiento #2', class MTA, trigger "Rec19" bit 11
   46: 'El Compresor ABC5 alcanzó la máxima cantidad de horas sin mantenimiento #2', class MTA, trigger "Rec19" bit 12
   47: 'El Compresor ABC1 alcanzó la máxima cantidad de horas sin mantenimiento #2', class MTA, trigger "Rec19" bit 13
   48: 'El Secador ABC1 superó la máxima cantidad de horas sin mantenimiento', class MTA, trigger "Rec20" bit 8
   49: 'El Secador ABC3 superó la máxima cantidad de horas sin mantenimiento', class MTA, trigger "Rec20" bit 9
   51: 'El Secador ABC2 superó la máxima cantidad de horas sin mantenimiento', class MTA, trigger "Rec20" bit 10
   52: 'El Secador Fargon superó la máxima cantidad de horas sin mantenimiento', class MTA, trigger "Rec20" bit 11
   54: 'El Secador Sullair 1 superó la máxima cantidad de horas sin mantenimiento #1', class MTA, trigger "Rec20" bit 12
   55: 'El Secador Sullair 1 superó la máxima cantidad de horas sin mantenimiento #2', class MTA, trigger "Rec20" bit 13
   56: 'El Secador Sullair 2 superó la máxima cantidad de horas sin mantenimiento #1', class MTA, trigger "Rec20" bit 14
   57: 'El Secador Sullair 2 superó la máxima cantidad de horas sin mantenimiento #2', class MTA, trigger "Rec20" bit 15
   58: 'El compresor Sullair 2 superó la máxima cantidad de horas sin mantenimiento #1', class MTA, trigger "Rec21" bit 8
   59: 'El compresor Sullair 2 superó la máxima cantidad de horas sin mantenimiento #2', class MTA, trigger "Rec21" bit 9
   60: 'El compresor Sullair 2 superó la máxima cantidad de horas sin mantenimiento #3', class MTA, trigger "Rec21" bit 10
   61: 'El compresor Sullair 2 superó la máxima cantidad de horas sin mantenimiento #4', class MTA, trigger "Rec21" bit 11
   62: 'El compresor Sullair 2 superó la máxima cantidad de horas sin mantenimiento #5', class MTA, trigger "Rec21" bit 12